       // Matching to PathData
       #parameterDefinition.directValues.cmdType := 3; // Circ Absolute
       #parameterDefinition.directValues.cmdParameters.circleParameters.circlePlane := 2; // XY
       #parameterDefinition.directValues.cmdParameters.circleParameters.pathChoice := 1; // neg rotation
       #parameterDefinition.directValues.cmdParameters.circleParameters.circMode := 3; // aux point is center relativ to start


     #G3:  // Circ CCW --> CircMode 1/2/3
       // Command name definition
       #parameterDefinition.parameterNameString := 'G';
       #parameterDefinition.parameterNameNumber := 3;

       // Properties
       #parameterDefinition.properties := "LKINLANG_MOTION_CMD" + "LKINLANG_CMD_MODAL";
       #parameterDefinition.validCountPerLine := 1;

       // Conditions
       #tempConditionCounter := 1;
       #parameterDefinition.conditions[#tempConditionCounter].ParameterNumber := #G17;
       #parameterDefinition.conditions[#tempConditionCounter].Group := 20;
       #parameterDefinition.conditions[#tempConditionCounter].Mode := "LKINLANG_CONDITION_IN_PROGRAM"; // In program
       #tempConditionCounter += 1;
       #parameterDefinition.conditions[#tempConditionCounter].ParameterNumber := #G18;
       #parameterDefinition.conditions[#tempConditionCounter].Group := 20;
       #parameterDefinition.conditions[#tempConditionCounter].Mode := "LKINLANG_CONDITION_IN_PROGRAM"; // In program
       #tempConditionCounter += 1;
       #parameterDefinition.conditions[#tempConditionCounter].ParameterNumber := #G19;
       #parameterDefinition.conditions[#tempConditionCounter].Group := 20;
       #parameterDefinition.conditions[#tempConditionCounter].Mode := "LKINLANG_CONDITION_IN_PROGRAM"; // In program
       #tempConditionCounter += 1;
       #parameterDefinition.conditions[#tempConditionCounter].ParameterNumber := #F;
       #parameterDefinition.conditions[#tempConditionCounter].Group := 10;
       #parameterDefinition.conditions[#tempConditionCounter].Mode := "LKINLANG_CONDITION_IN_PROGRAM"; // In program

       // Priorities
       // PathChoice and CmdType are defined
       #parameterDefinition.priorities.cmdType := "LKINLANG_PRIO_DEFINED";
       #parameterDefinition.priorities.cmdParameters.circleParameters.pathChoice := "LKINLANG_PRIO_DEFINED";

       // CircMode and circPlane can be changed (G17,G18,G19 / AR,CR,I,J,K)
       #parameterDefinition.priorities.cmdParameters.circleParameters.circlePlane := "LKINLANG_PRIO_DEFAULT";
       #parameterDefinition.priorities.cmdParameters.circleParameters.circMode := "LKINLANG_PRIO_DEFAULT";

       // Matching to PathData
       #parameterDefinition.directValues.cmdType := 3;
       #parameterDefinition.directValues.cmdParameters.circleParameters.circlePlane := 2; // XY
       #parameterDefinition.directValues.cmdParameters.circleParameters.pathChoice := 0; // pos rotation
       #parameterDefinition.directValues.cmdParameters.circleParameters.circMode := 3; // aux point is center relativ to start

     #G5:  // Circ 3D --> CircMode 0 
       // Command name definition
       #parameterDefinition.parameterNameString := 'G';
       #parameterDefinition.parameterNameNumber := 5;

       // Properties
       #parameterDefinition.properties := "LKINLANG_MOTION_CMD" + "LKINLANG_CMD_MODAL";
       #parameterDefinition.validCountPerLine := 1;

       // Conditions
       #tempConditionCounter := 1;
       #parameterDefinition.conditions[#tempConditionCounter].ParameterNumber := #F;
       #parameterDefinition.conditions[#tempConditionCounter].Group := 10;
       #parameterDefinition.conditions[#tempConditionCounter].Mode := "LKINLANG_CONDITION_IN_PROGRAM"; // In program

       // Priorities
       // CmdType and CircMode are defined 
       #parameterDefinition.priorities.cmdType := "LKINLANG_PRIO_DEFINED";
       #parameterDefinition.priorities.cmdParameters.circleParameters.circMode := "LKINLANG_PRIO_DEFINED";

       // Matching to PathData
       #parameterDefinition.directValues.cmdType := 3;
       #parameterDefinition.directValues.cmdParameters.circleParameters.circMode := 0; // aux point is on circ line


     #G4: // Wait time
       // Command name definition
       #parameterDefinition.parameterNameString := 'G';
       #parameterDefinition.parameterNameNumber := 4;

       // Properties
       #parameterDefinition.properties := 16#0;//"LKINLANG_MOTION_CMD";
       #parameterDefinition.validCountPerLine := 1;

       // Conditions
       #tempConditionCounter := 1;
       #parameterDefinition.conditions[#tempConditionCounter].ParameterNumber := #P;
       #parameterDefinition.conditions[#tempConditionCounter].Group := 30;
       #parameterDefinition.conditions[#tempConditionCounter].Mode := "LKINLANG_CONDITION_IN_LINE"; // In line

       #tempConditionCounter += 1;
       #parameterDefinition.conditions[#tempConditionCounter].ParameterNumber := #F;
       #parameterDefinition.conditions[#tempConditionCounter].Group := 30;
       #parameterDefinition.conditions[#tempConditionCounter].Mode := "LKINLANG_CONDITION_IN_LINE"; // In line

       // Properties
       #parameterDefinition.priorities.cmdType := "LKINLANG_PRIO_DEFINED";

       // Matching to PathData
       #parameterDefinition.directValues.cmdType := 100;

     #P: // WaitTime, same as F?
       // Command name definition
       #parameterDefinition.parameterNameString := 'P';
       #parameterDefinition.parameterNameNumber := -1;

       // Properties
       #parameterDefinition.properties := "LKINLANG_EQUATION";
       #parameterDefinition.validCountPerLine := 1;

       // Priorities
       #parameterDefinition.priorities.cmdParameters.pathDynamics.velocity := "LKINLANG_PRIO_DEFINED";

       // Matching to PathData
       #parameterDefinition.followingValues[1].cmdParameters.pathDynamics.velocity := TRUE;


     #G40: // Tool off
       // Command name definition
       #parameterDefinition.parameterNameString := 'G';
       #parameterDefinition.parameterNameNumber := 40;

       // Properties
       #parameterDefinition.properties := 16#0;//"LKINLANG_MOTION_CMD";

       // Priorities
       #parameterDefinition.priorities.cmdType := "LKINLANG_PRIO_DEFINED";

       // Matching to PathData
       #parameterDefinition.directValues.cmdType := 40;

     #G41: // Tool left
       // Command name definition
       #parameterDefinition.parameterNameString := 'G';
       #parameterDefinition.parameterNameNumber := 41;

       // Properties
       #parameterDefinition.properties := 16#0;//"LKINLANG_MOTION_CMD";

       // Priorities
       #parameterDefinition.priorities.cmdType := "LKINLANG_PRIO_DEFINED";

       // Matching to PathData
       #parameterDefinition.directValues.cmdType := 41;

       // Conditions
       #tempConditionCounter := 1;
       #parameterDefinition.conditions[#tempConditionCounter].ParameterNumber := #T;
       #parameterDefinition.conditions[#tempConditionCounter].Group := 40;
       #parameterDefinition.conditions[#tempConditionCounter].Mode := "LKINLANG_CONDITION_IN_PROGRAM";
       #tempConditionCounter += 1;
       #parameterDefinition.conditions[#tempConditionCounter].ParameterNumber := #G17;
       #parameterDefinition.conditions[#tempConditionCounter].Group := 20;
       #parameterDefinition.conditions[#tempConditionCounter].Mode := "LKINLANG_CONDITION_IN_PROGRAM"; // In program
       #tempConditionCounter += 1;
       #parameterDefinition.conditions[#tempConditionCounter].ParameterNumber := #G18;
       #parameterDefinition.conditions[#tempConditionCounter].Group := 20;
       #parameterDefinition.conditions[#tempConditionCounter].Mode := "LKINLANG_CONDITION_IN_PROGRAM"; // In program
       #tempConditionCounter += 1;
       #parameterDefinition.conditions[#tempConditionCounter].ParameterNumber := #G19;
       #parameterDefinition.conditions[#tempConditionCounter].Group := 20;
       #parameterDefinition.conditions[#tempConditionCounter].Mode := "LKINLANG_CONDITION_IN_PROGRAM"; // In program

     #G42: // Tool right
       // Command name definition
       #parameterDefinition.parameterNameString := 'G';
       #parameterDefinition.parameterNameNumber := 42;

       // Properties
       #parameterDefinition.properties := 16#0; //"LKINLANG_MOTION_CMD";

       // Priorities
       #parameterDefinition.priorities.cmdType := "LKINLANG_PRIO_DEFINED";

       // Matching to PathData
       #parameterDefinition.directValues.cmdType := 42;

       // Conditions
       #tempConditionCounter := 1;
       #parameterDefinition.conditions[#tempConditionCounter].ParameterNumber := #T;
       #parameterDefinition.conditions[#tempConditionCounter].Group := 40;
       #parameterDefinition.conditions[#tempConditionCounter].Mode := "LKINLANG_CONDITION_IN_PROGRAM";
       #tempConditionCounter += 1;
       #parameterDefinition.conditions[#tempConditionCounter].ParameterNumber := #G17;
       #parameterDefinition.conditions[#tempConditionCounter].Group := 20;
       #parameterDefinition.conditions[#tempConditionCounter].Mode := "LKINLANG_CONDITION_IN_PROGRAM"; // In program
       #tempConditionCounter += 1;
       #parameterDefinition.conditions[#tempConditionCounter].ParameterNumber := #G18;
       #parameterDefinition.conditions[#tempConditionCounter].Group := 20;
       #parameterDefinition.conditions[#tempConditionCounter].Mode := "LKINLANG_CONDITION_IN_PROGRAM"; // In program
       #tempConditionCounter += 1;
       #parameterDefinition.conditions[#tempConditionCounter].ParameterNumber := #G19;
       #parameterDefinition.conditions[#tempConditionCounter].Group := 20;
       #parameterDefinition.conditions[#tempConditionCounter].Mode := "LKINLANG_CONDITION_IN_PROGRAM"; // In program

     #T: // Tool selection
       // Command name definition
       #parameterDefinition.parameterNameString := 'T';
       #parameterDefinition.parameterNameNumber := -1;

       #parameterDefinition.validCountPerLine := 1;

       // Properties
       #parameterDefinition.properties := "LKINLANG_PRG_MODAL";

       // Matching to PathData
       #parameterDefinition.priorities.cmdParameters.offsetParameters.offsetParaNo := "LKINLANG_PRIO_DEFINED";
       #parameterDefinition.followingValues[1].cmdParameters.offsetParameters.offsetParaNo := TRUE;


     #G17: // XY PathPlane
       // Command name definition
       #parameterDefinition.parameterNameString := 'G';
       #parameterDefinition.parameterNameNumber := 17;

       // Properties
       #parameterDefinition.properties := "LKINLANG_PRG_MODAL";

       // Matching to PathData
       #parameterDefinition.priorities.cmdParameters.circleParameters.circlePlane := "LKINLANG_PRIO_DEFINED";
       #parameterDefinition.directValues.cmdParameters.circleParameters.circlePlane := 2; // XY

       // Also set main path plane
       #parameterDefinition.priorities.cmdParameters.offsetParameters.mainPathPlane := "LKINLANG_PRIO_DEFINED";
       #parameterDefinition.directValues.cmdParameters.offsetParameters.mainPathPlane := 2; // XY

     #G18: // XZ PathPlane
       // Command name definition
       #parameterDefinition.parameterNameString := 'G';
       #parameterDefinition.parameterNameNumber := 18;

       // Properties
       #parameterDefinition.properties := "LKINLANG_PRG_MODAL";

       // Matching to PathData
       #parameterDefinition.priorities.cmdParameters.circleParameters.circlePlane := "LKINLANG_PRIO_DEFINED";
       #parameterDefinition.directValues.cmdParameters.circleParameters.circlePlane := 0; // XZ

       // Also set main path plane
       #parameterDefinition.priorities.cmdParameters.offsetParameters.mainPathPlane := "LKINLANG_PRIO_DEFINED";
       #parameterDefinition.directValues.cmdParameters.offsetParameters.mainPathPlane := 0; // XZ

     #G19: //YZ PathPlane
       // Command name definition
       #parameterDefinition.parameterNameString := 'G';
       #parameterDefinition.parameterNameNumber := 19;

       // Properties
       #parameterDefinition.properties := "LKINLANG_PRG_MODAL";

       // Matching to PathData
       #parameterDefinition.priorities.cmdParameters.circleParameters.circlePlane := "LKINLANG_PRIO_DEFINED";
       #parameterDefinition.directValues.cmdParameters.circleParameters.circlePlane := 1; // YZ

       // Also set main path plane
       #parameterDefinition.priorities.cmdParameters.offsetParameters.mainPathPlane := "LKINLANG_PRIO_DEFINED";
       #parameterDefinition.directValues.cmdParameters.offsetParameters.mainPathPlane := 1; // YZ

     #G640:
       // Command name definition
       #parameterDefinition.parameterNameString := 'G';
       #parameterDefinition.parameterNameNumber := 640;

       // Properties
       #parameterDefinition.properties := "LKINLANG_PRG_MODAL";

       // Matching to PathData
       #parameterDefinition.priorities.cmdParameters.bufferMode := "LKINLANG_PRIO_DEFINED";
       #parameterDefinition.directValues.cmdParameters.bufferMode := 1; // Standstill

       #parameterDefinition.priorities.cmdParameters.transitionParameters[1] := "LKINLANG_PRIO_DEFINED";
       #parameterDefinition.directValues.cmdParameters.transitionParameters[1] := 0.0; // Standstill

     #G641:
       // Command name definition
       #parameterDefinition.parameterNameString := 'G';
       #parameterDefinition.parameterNameNumber := 641;

       // Properties
       #parameterDefinition.properties := "LKINLANG_PRG_MODAL";

       // Conditions
       #tempConditionCounter := 1;
       #parameterDefinition.conditions[#tempConditionCounter].ParameterNumber := #BR;
       #parameterDefinition.conditions[#tempConditionCounter].Group := 50;
       #parameterDefinition.conditions[#tempConditionCounter].Mode := "LKINLANG_CONDITION_IN_LINE"; // In line

       // Matching to PathData
       #parameterDefinition.priorities.cmdParameters.bufferMode := "LKINLANG_PRIO_DEFINED";
       #parameterDefinition.directValues.cmdParameters.bufferMode := #parameterDefaults.transitionVelocityMode;

     #G90:
       // Command name definition
       #parameterDefinition.parameterNameString := 'G';
       #parameterDefinition.parameterNameNumber := 90;

       // Properties
       #parameterDefinition.properties := "LKINLANG_PRG_MODAL" + "LKINLANG_ABSOLUTE_POSITION";


     #G91:
       // Command name definition
       #parameterDefinition.parameterNameString := 'G';
       #parameterDefinition.parameterNameNumber := 91;

       // Properties
       #parameterDefinition.properties := "LKINLANG_PRG_MODAL" + "LKINLANG_RELATIVE_POSITION";

     #G54: // Select OCS 1
       // Command name definition
       #parameterDefinition.parameterNameString := 'G';
       #parameterDefinition.parameterNameNumber := 54;

       // Properties
       #parameterDefinition.properties := "LKINLANG_PRG_MODAL" + "LKINLANG_CHECK_LIMITS";

       // Matching to PathData
       #parameterDefinition.priorities.cmdCoordinates.coordSystem := "LKINLANG_PRIO_DEFINED";
       #parameterDefinition.directValues.cmdCoordinates.coordSystem := 1; // OCS1


     #G55: // Select OCS 2
       // Command name definition
       #parameterDefinition.parameterNameString := 'G';
       #parameterDefinition.parameterNameNumber := 55;

       // Properties
       #parameterDefinition.properties := "LKINLANG_PRG_MODAL" + "LKINLANG_CHECK_LIMITS";

       // Matching to PathData
       #parameterDefinition.priorities.cmdCoordinates.coordSystem := "LKINLANG_PRIO_DEFINED";
       #parameterDefinition.directValues.cmdCoordinates.coordSystem := 2; // OCS2


     #G56: // Select OCS 3
       // Command name definition
       #parameterDefinition.parameterNameString := 'G';
       #parameterDefinition.parameterNameNumber := 56;

       // Properties
       #parameterDefinition.properties := "LKINLANG_PRG_MODAL" + "LKINLANG_CHECK_LIMITS";

       // Matching to PathData
       #parameterDefinition.priorities.cmdCoordinates.coordSystem := "LKINLANG_PRIO_DEFINED";
       #parameterDefinition.directValues.cmdCoordinates.coordSystem := 3; // OCS3


     #G500: // Select WCS
       // Command name definition
       #parameterDefinition.parameterNameString := 'G';
       #parameterDefinition.parameterNameNumber := 500;

       // Properties
       #parameterDefinition.properties := "LKINLANG_PRG_MODAL" + "LKINLANG_CHECK_LIMITS";

       // Matching to PathData
       #parameterDefinition.priorities.cmdCoordinates.coordSystem := "LKINLANG_PRIO_DEFINED";
       #parameterDefinition.directValues.cmdCoordinates.coordSystem := 0; // WCS


       // Gerneral Parameters (170 - 199)
       // ===========================================================
     #X:
       #parameterDefinition.parameterNameString := 'X';
       #parameterDefinition.parameterNameNumber := -1;
       #parameterDefinition.properties := "LKINLANG_CHECK_LIMITS" + "LKINLANG_EQUATION";
       #parameterDefinition.priorities.cmdCoordinates.cartesianPosition.x := "LKINLANG_PRIO_DEFINED";
       #parameterDefinition.followingValues[1].cmdCoordinates.cartesianPosition.x := true;

     #Y:
       #parameterDefinition.parameterNameString := 'Y';
       #parameterDefinition.parameterNameNumber := -1;
       #parameterDefinition.properties := "LKINLANG_CHECK_LIMITS" + "LKINLANG_EQUATION";
       #parameterDefinition.priorities.cmdCoordinates.cartesianPosition.y := "LKINLANG_PRIO_DEFINED";
       #parameterDefinition.followingValues[1].cmdCoordinates.cartesianPosition.y := true;

     #Z:
       #parameterDefinition.parameterNameString := 'Z';
       #parameterDefinition.parameterNameNumber := -1;
       #parameterDefinition.properties := "LKINLANG_CHECK_LIMITS" + "LKINLANG_EQUATION";
       #parameterDefinition.priorities.cmdCoordinates.cartesianPosition.z := "LKINLANG_PRIO_DEFINED";
       #parameterDefinition.followingValues[1].cmdCoordinates.cartesianPosition.z := true;

     #A:
       #parameterDefinition.parameterNameString := 'A';
       #parameterDefinition.parameterNameNumber := -1;
       #parameterDefinition.properties := "LKINLANG_CHECK_LIMITS" + "LKINLANG_EQUATION";
       #parameterDefinition.priorities.cmdCoordinates.cartesianPosition.a := "LKINLANG_PRIO_DEFINED";
       #parameterDefinition.followingValues[1].cmdCoordinates.cartesianPosition.a := true;

       // Orientation direction
       #parameterDefinition.directValues.cmdParameters.orientationDirection := #parameterDefaults.orientationDirection;
       #parameterDefinition.directValues.cmdParameters.orientationDirection := "LKINLANG_PRIO_DEFAULT";

     #F:
       #parameterDefinition.parameterNameString := 'F';
       #parameterDefinition.parameterNameNumber := -1;
       #parameterDefinition.properties := "LKINLANG_PRG_MODAL" + "LKINLANG_CHECK_LIMITS" + "LKINLANG_EQUATION";
       #parameterDefinition.priorities.cmdParameters.pathDynamics.velocity := "LKINLANG_PRIO_DEFINED";
       #parameterDefinition.followingValues[1].cmdParameters.pathDynamics.velocity := TRUE;

     #ACC:
       #parameterDefinition.parameterNameString := 'ACC';
       #parameterDefinition.parameterNameNumber := -1;
       #parameterDefinition.properties := "LKINLANG_PRG_MODAL" + "LKINLANG_CHECK_LIMITS" + "LKINLANG_EQUATION";
       #parameterDefinition.priorities.cmdParameters.pathDynamics.acceleration := "LKINLANG_PRIO_DEFINED";
       #parameterDefinition.followingValues[1].cmdParameters.pathDynamics.acceleration := TRUE;

     #DEC:
       #parameterDefinition.parameterNameString := 'DEC';
       #parameterDefinition.parameterNameNumber := -1;
       #parameterDefinition.properties := "LKINLANG_PRG_MODAL" + "LKINLANG_CHECK_LIMITS" + "LKINLANG_EQUATION";
       #parameterDefinition.priorities.cmdParameters.pathDynamics.deceleration := "LKINLANG_PRIO_DEFINED";
       #parameterDefinition.followingValues[1].cmdParameters.pathDynamics.deceleration := TRUE;

     #JERK:
       #parameterDefinition.parameterNameString := 'JERK';
       #parameterDefinition.parameterNameNumber := -1;
       #parameterDefinition.properties := "LKINLANG_PRG_MODAL" + "LKINLANG_CHECK_LIMITS" + "LKINLANG_EQUATION";
       #parameterDefinition.priorities.cmdParameters.pathDynamics.jerk := "LKINLANG_PRIO_DEFINED";
       #parameterDefinition.followingValues[1].cmdParameters.pathDynamics.jerk := TRUE;


     #I:
       // Command name definition
       #parameterDefinition.parameterNameString := 'I';
       #parameterDefinition.parameterNameNumber := -1;

       // Properties
       #parameterDefinition.properties := "LKINLANG_EQUATION";

       // Matching to PathData
       #parameterDefinition.priorities.cmdParameters.circleParameters.auxPoint[1] := "LKINLANG_PRIO_DEFINED";
       #parameterDefinition.followingValues[1].cmdParameters.circleParameters.auxPoint[1] := TRUE;

     #J:
       // Command name definition
       #parameterDefinition.parameterNameString := 'J';
       #parameterDefinition.parameterNameNumber := -1;

       // Properties
       #parameterDefinition.properties := "LKINLANG_EQUATION";

       // Matching to PathData
       #parameterDefinition.priorities.cmdParameters.circleParameters.auxPoint[2] := "LKINLANG_PRIO_DEFINED";
       #parameterDefinition.followingValues[1].cmdParameters.circleParameters.auxPoint[2] := TRUE;

     #K:
       // Command name definition
       #parameterDefinition.parameterNameString := 'K';
       #parameterDefinition.parameterNameNumber := -1;

       // Properties
       #parameterDefinition.properties := "LKINLANG_EQUATION";

       // Matching to PathData
       #parameterDefinition.priorities.cmdParameters.circleParameters.auxPoint[3] := "LKINLANG_PRIO_DEFINED";
       #parameterDefinition.followingValues[1].cmdParameters.circleParameters.auxPoint[3] := TRUE;

     #AR:
       // Command name definition
       #parameterDefinition.parameterNameString := 'AR';
       #parameterDefinition.parameterNameNumber := -1;

       // Properties
       #parameterDefinition.properties := "LKINLANG_EQUATION";

       // Conditions
       #tempConditionCounter := 1;
       #parameterDefinition.conditions[#tempConditionCounter].ParameterNumber := #I;
       #parameterDefinition.conditions[#tempConditionCounter].Group := 60;
       #parameterDefinition.conditions[#tempConditionCounter].Mode := "LKINLANG_CONDITION_IN_LINE"; // In Line
       #tempConditionCounter += 1; 
       #parameterDefinition.conditions[#tempConditionCounter].ParameterNumber := #J;
       #parameterDefinition.conditions[#tempConditionCounter].Group := 60;
       #parameterDefinition.conditions[#tempConditionCounter].Mode := "LKINLANG_CONDITION_IN_LINE"; // In Line
       #tempConditionCounter += 1;
       #parameterDefinition.conditions[#tempConditionCounter].ParameterNumber := #K;
       #parameterDefinition.conditions[#tempConditionCounter].Group := 60;
       #parameterDefinition.conditions[#tempConditionCounter].Mode := "LKINLANG_CONDITION_IN_LINE"; // In Line

       // Matching to PathData
       #parameterDefinition.priorities.cmdParameters.circleParameters.arc := "LKINLANG_PRIO_DEFINED";
       #parameterDefinition.followingValues[1].cmdParameters.circleParameters.arc := TRUE;
       #parameterDefinition.priorities.cmdParameters.circleParameters.circMode := "LKINLANG_PRIO_DEFINED";
       #parameterDefinition.directValues.cmdParameters.circleParameters.circMode := 1;

     #CR:
       // Command name definition
       #parameterDefinition.parameterNameString := 'CR';
       #parameterDefinition.parameterNameNumber := -1;

       // Properties
       #parameterDefinition.properties := "LKINLANG_EQUATION";

       // Conditions
       #tempConditionCounter := 1;
       #parameterDefinition.conditions[#tempConditionCounter].ParameterNumber := #X;
       #parameterDefinition.conditions[#tempConditionCounter].Group := 70;
       #parameterDefinition.conditions[#tempConditionCounter].Mode := "LKINLANG_CONDITION_IN_LINE"; // In Line
       #tempConditionCounter += 1;
       #parameterDefinition.conditions[#tempConditionCounter].ParameterNumber := #Y;
       #parameterDefinition.conditions[#tempConditionCounter].Group := 70;
       #parameterDefinition.conditions[#tempConditionCounter].Mode := "LKINLANG_CONDITION_IN_LINE"; // In Line
       #tempConditionCounter += 1;
       #parameterDefinition.conditions[#tempConditionCounter].ParameterNumber := #Z;
       #parameterDefinition.conditions[#tempConditionCounter].Group := 70;
       #parameterDefinition.conditions[#tempConditionCounter].Mode := "LKINLANG_CONDITION_IN_LINE"; // In Line

       // Matching to PathData
       #parameterDefinition.priorities.cmdParameters.circleParameters.radius := "LKINLANG_PRIO_DEFINED";
       #parameterDefinition.followingValues[1].cmdParameters.circleParameters.radius := TRUE;
       #parameterDefinition.priorities.cmdParameters.circleParameters.circMode := "LKINLANG_PRIO_DEFINED";
       #parameterDefinition.directValues.cmdParameters.circleParameters.circMode := 2;

     #M:
       // Command name definition
       #parameterDefinition.parameterNameString := 'M';
       #parameterDefinition.parameterNameNumber := -1;

       #parameterDefinition.validCountPerLine := "LKINCTRL_NO_OF_CMD_SETFLAGS";

       // Properties
       #parameterDefinition.properties := "LKINLANG_CHECK_LIMITS";

       // Matching to PathData
       #parameterDefinition.priorities.setFlags.flag := "LKINLANG_PRIO_DEFINED";
       #parameterDefinition.priorities.setFlags.flagMode := "LKINLANG_PRIO_DEFINED";
       #parameterDefinition.priorities.setFlags.remainingDistance := "LKINLANG_PRIO_DEFINED";
       #parameterDefinition.followingValues[1].setFlags.flag := TRUE;
       #parameterDefinition.followingValues[2].setFlags.flagMode := TRUE;
       #parameterDefinition.followingValues[3].setFlags.remainingDistance := TRUE;

     #H:
       // Command name definition
       #parameterDefinition.parameterNameString := 'H';
       #parameterDefinition.parameterNameNumber := -1;

       #parameterDefinition.validCountPerLine := "LKINCTRL_NO_OF_CMD_SETFLAGS";

       // Properties
       #parameterDefinition.properties := "LKINLANG_CHECK_LIMITS" + "LKINLANG_EQUATION";

       // Matching to PathData
       #parameterDefinition.priorities.valueFlags.flag := "LKINLANG_PRIO_DEFINED";
       #parameterDefinition.priorities.valueFlags.value := "LKINLANG_PRIO_DEFINED";
       #parameterDefinition.priorities.valueFlags.flagMode := "LKINLANG_PRIO_DEFINED";
       #parameterDefinition.priorities.valueFlags.remainingDistance := "LKINLANG_PRIO_DEFINED";
       #parameterDefinition.followingValues[1].valueFlags.flag := TRUE;
       #parameterDefinition.followingValues[2].valueFlags.value := TRUE;
       #parameterDefinition.followingValues[3].valueFlags.flagMode := TRUE;
       #parameterDefinition.followingValues[4].valueFlags.remainingDistance := TRUE;

     #BR:
       // Command name definition
       #parameterDefinition.parameterNameString := 'BR';
       #parameterDefinition.parameterNameNumber := -1;

       // Properties
       #parameterDefinition.properties := "LKINLANG_PRG_MODAL" + "LKINLANG_EQUATION";

       // Matching to PathData
       #parameterDefinition.priorities.cmdParameters.transitionParameters[1] := "LKINLANG_PRIO_DEFINED";
       #parameterDefinition.followingValues[1].cmdParameters.transitionParameters[1] := TRUE;

     #M30:
       // Command name definition
       #parameterDefinition.parameterNameString := 'M';
       #parameterDefinition.parameterNameNumber := 30;

       #parameterDefinition.validCountPerLine := 1;

       // Properties
       #parameterDefinition.properties := "LKINLANG_MOTION_CMD";
       #parameterDefinition.priorities.cmdType := "LKINLANG_PRIO_DEFINED";

       // Matching to PathData
       #parameterDefinition.directValues.cmdType := -1;
     ELSE
       // invalid case number
       #parameterNo := -2;

   END_CASE;
END_FUNCTION

FUNCTION "LKinLang_UserDefinedGCode" : Void   // FC35453, SCL
TITLE = LKinLang_LangPackageGCode
{ S7_Optimized_Access := 'TRUE' }
AUTHOR : tech.team.motioncontrol@siemens.com
FAMILY : LKinLang
VERSION : 1.1
// Language definition package for user defined GCode
   VAR_IN_OUT
      parameterNo : Int;   // Parameter number
      parameterDefinition : "LKinLang_typeParameterDefinition";   // Found parameter definition
      parameterDefaults : "LKinLang_typeGCodeDefaults";   // Parameter defaults
   END_VAR
   VAR_TEMP
      tempConditionCounter : Int;
   END_VAR
   VAR CONSTANT
      G0 : DInt := 100;   // Fast Lin
      G1 : DInt := 101;   // Lin
      G2 : DInt := 102;   // Circ CW
      G3 : DInt := 103;   // Circ CCW
      G5 : DInt := 105;   // Circ 3D
      G4 : DInt := 104;   // WaitTime
      P : DInt := 110;   // Period for WaitTime
      G17 : DInt := 120;   // XY Plane
      G18 : DInt := 121;   // ZX Plane
      G19 : DInt := 122;   // YZ Plane
      G640 : DInt := 130;   // Geometry blending off
      G641 : DInt := 131;   // Geometry blending with high velocity
      G642 : DInt := 132;   // Geometry blending with low velocity
      G90 : DInt := 150;   // Absolute Position
      G91 : DInt := 151;   // Relativ Position
      G54 : DInt := 152;   // Select OCS1
      G55 : DInt := 153;   // Select OCS2
      G56 : DInt := 154;   // Select OCS3
      G500 : DInt := 155;   // Select WCS
      T : DInt := 160;   // Tool selection
      G40 : DInt := 161;   // Tool off
      G41 : DInt := 162;   // Tool left
      G42 : DInt := 163;   // Tool right
      X : DInt := 170;   // X pos
      Y : DInt := 171;   // Y pos
      Z : DInt := 172;   // Z pos
      "A" : DInt := 173;   // Orientation
      F : DInt := 174;   // Velocity
      ACC : DInt := 175;   // Acceleration
      DEC : DInt := 176;   // Deceleration
      JERK : DInt := 177;   // Jerk
      CR : DInt := 178;   // Circle Radius
      I : DInt := 179;   // Circ Point
      J : DInt := 180;   // Circ Point
      K : DInt := 181;   // Circ Point
      AR : DInt := 182;   // Arc
      BR : DInt := 183;   // Transition Parameter
      "M" : DInt := 190;   // Flag
      M30 : DInt := 199;   // End of PRG
   END_VAR
BEGIN
   //==========================================================================================
   // SIEMENS AG
   // (c)Copyright 2019 All Rights Reserved
   //------------------------------------------------------------------------------------------
   // Library: LKinLang
   // Tested with: S7-1517T-3 PN/DP
   // Engineering: TIA Portal V15
   // Restrictions: ---
   // Requirements: S7-1500T FW 2.5
   // Functionality: LKinLang_UserDefinedGCode
   // Language definition package for user defined GCode
   // 
   // Support: tech.team.motioncontrol@siemens.com
   // Note: Parameter comments are only available in language 'English (United States)'
   //------------------------------------------------------------------------------------------
   // Change log table:
   // Version    Date          Expert in charge    Changes applied
   // 01.00.00   28.05.2019    FR                  First created version
   //===========================================================================================
   //
   //  Group Parameter 
   //  10:   F
   //        
   //  20:   G17
   //        G18
   //        G19
   //        
   //  30:   F
   //        P
   //        
   //  40:   T
   //
   //  50:   BR
   //  
   //  60:   I
   //        J
   //        K
   //
   //  70:   X
   //        Y
   //        Z


   CASE #parameterNo OF
       // User defined commands for GCode.
       // Here you can define up to 100 commands.
       // It is possible to overload predefined GCode commands.
       // Or define own commands.
       // Some example are already programmed.
       // ------------------------------
     1:
       // ========================================================================================================
       // End of program
       // ========================================================================================================
       // Instead of M30, END is also possible
       // ========================================================================================================
       // Parameter name definition
       #parameterDefinition.parameterNameString := 'END';
       #parameterDefinition.parameterNameNumber := -1;

       // Matching to PathData
       #parameterDefinition.directValues.cmdType := -1;

       // Priorities
       #parameterDefinition.priorities.cmdType := "LKINLANG_PRIO_DEFINED";

       // Properties
       #parameterDefinition.properties := "LKINLANG_MOTION_CMD";

       // Valid counts per line
       #parameterDefinition.validCountPerLine := 1;
       // ========================================================================================================

     2:
       // ========================================================================================================
       // Gripper control ON
       // ========================================================================================================
       // This is an example for an defined "Gripper" parameter
       // 'GRIPPER_ON' sets Flag 1 with Flagmode 11
       // ========================================================================================================
       // Parameter name definition
       #parameterDefinition.parameterNameString := 'GRIPPER_ON';
       #parameterDefinition.parameterNameNumber := -1;

       // Matching to PathData
       #parameterDefinition.directValues.setFlags[1].flag := 1;
       #parameterDefinition.directValues.setFlags[1].flagMode := 11;

       // Priorities
       #parameterDefinition.priorities.setFlags.flag := "LKINLANG_PRIO_DEFINED";
       #parameterDefinition.priorities.setFlags.flagMode := "LKINLANG_PRIO_DEFINED";

       // Properties
       #parameterDefinition.properties := 16#0;

       // Valid counts per line
       #parameterDefinition.validCountPerLine := 1;
       // ========================================================================================================

     3:
       // ========================================================================================================
       // Gripper control OFF
       // ========================================================================================================
       // This is an example for an defined "Gripper" parameter
       // 'GRIPPER_OFF' resets Flag 1 with Flagmode 13
       // ========================================================================================================
       // Parameter name definition
       #parameterDefinition.parameterNameString := 'GRIPPER_OFF';
       #parameterDefinition.parameterNameNumber := -1;

       // Matching to PathData
       #parameterDefinition.directValues.setFlags[1].flag := 1;
       #parameterDefinition.directValues.setFlags[1].flagMode := 13;

       // Priorities
       #parameterDefinition.priorities.setFlags.flag := "LKINLANG_PRIO_DEFINED";
       #parameterDefinition.priorities.setFlags.flagMode := "LKINLANG_PRIO_DEFINED";

       // Properties
       #parameterDefinition.properties := 16#0;

       // Valid counts per line
       #parameterDefinition.validCountPerLine := 1;
       // ========================================================================================================

     4: 
       // ========================================================================================================
       // Point name
       // ========================================================================================================
       // Use 'Nxx' as point name in the PathData
       // --> Only numbers possible
       // ========================================================================================================
       // Parameter name definition
       #parameterDefinition.parameterNameString := 'N';
       #parameterDefinition.parameterNameNumber := -1;

       // Matching to PathData
       #parameterDefinition.followingValues[1].cmdName := TRUE;

       // Priorities
       #parameterDefinition.priorities.cmdName := "LKINLANG_PRIO_DEFINED";

       // Properties
       #parameterDefinition.properties := 16#0;

       // Valid counts per line
       #parameterDefinition.validCountPerLine := 1;
       // ========================================================================================================

     5:
       // ========================================================================================================
       // Blending with low velocity
       // ========================================================================================================
       // Parameter name definition
       #parameterDefinition.parameterNameString := 'G';
       #parameterDefinition.parameterNameNumber := 642;

       // Matching to PathData
       #parameterDefinition.directValues.cmdParameters.bufferMode := 2; // Blending with low velocity

       // Priorites
       #parameterDefinition.priorities.cmdParameters.bufferMode := "LKINLANG_PRIO_DEFINED";

       // Properties
       #parameterDefinition.properties := "LKINLANG_PRG_MODAL";

       // Conditions
       #tempConditionCounter := 1;
       #parameterDefinition.conditions[#tempConditionCounter].ParameterNumber := #BR;
       #parameterDefinition.conditions[#tempConditionCounter].Group := 50;
       #parameterDefinition.conditions[#tempConditionCounter].Mode := "LKINLANG_CONDITION_IN_LINE"; // "BR" must be written in the same line

       // Valid counts per line
       #parameterDefinition.validCountPerLine := 1;
       // ========================================================================================================

     ELSE
       // invalid case number
       #parameterNo := -2;
   END_CASE;
END_FUNCTION

// folder: LKinLang_Blocks/LKinLang_LanguageDefinition/LKinLang_LangPackUser

FUNCTION "LKinLang_LangPackageUser" : Void   // FC35487, SCL
TITLE = LKinLang_LangPackageUser
{ S7_Optimized_Access := 'TRUE' }
AUTHOR : tech.team.motioncontrol@siemens.com
FAMILY : LKinLang
VERSION : 1.1
// Language definition package for a user defined language
   VAR_IN_OUT
      parameterNo : Int;   // Parameter number
      parameterDefinition : "LKinLang_typeParameterDefinition";   // Found parameter definition / Found command definition
      parameterDefaults : "LKinLang_typeUserDefinedDefaults";   // Parameter defaults
   END_VAR
   VAR_TEMP
      tempConditionCounter : Int;   // Temporary counter
   END_VAR
   VAR CONSTANT
      LIN : DInt := 1;   // Fast Lin
      VEL : DInt := 2;   // Velocity / Circ CW
      BLEND : DInt := 3;   // Blending
      RADIUS : DInt := 4;   // Blending radius
      X : DInt := 5;   // X pos
      Y : DInt := 6;   // Y pos
      Z : DInt := 7;   // Z pos
      END : DInt := 8;   // End of PRG
   END_VAR
BEGIN
   //==========================================================================================
   // SIEMENS AG
   // (c)Copyright 2019 All Rights Reserved
   //------------------------------------------------------------------------------------------
   // Library: LKinLang
   // Tested with: S7-1517T-3 PN/DP
   // Engineering: TIA Portal V15
   // Restrictions: ---
   // Requirements: S7-1500T FW 2.5
   // Functionality: LKinLang_LangPackageUser
   // Language definition package for completly user defined language
   // 
   // Support: tech.team.motioncontrol@siemens.com
   // Note: Parameter comments are only available in language 'English (United States)'
   //------------------------------------------------------------------------------------------
   // Change log table:
   // Version    Date          Expert in charge    Changes applied
   // 01.00.00   28.05.2019    FR                  First created version
   //===========================================================================================
   //
   //  Group Parameter 
   //  10:   R
   //        

   CASE #parameterNo OF
       // ========================================================================================================
       // Motion Parameters
       // ========================================================================================================
     #LIN:
       // ========================================================================================================
       // Linear movement
       // ========================================================================================================
       // Definition of linear movement (PathData: cmdType = 1) with default velocity
       // Parameter name is defined by parameterNameString and parameterNameNumber
       // ParameterNameString = LIN
       // ParameterNameNumber = -1 --> irrelevant
       // ==> Program line is searched for "LIN"

       // If "LIN" was found, set the defined values in the connected PathData.
       // The values are defined as "DirectValues" because the value to set is directly written here in this FC
       // Command type (cmdType)
       // #parameterDefinition.directValues.cmdType := 1;
       // --> Set the cmdType to 1
       // 
       // Velocity
       // #parameterDefinition.directValues.cmdParameters.pathDynamics.velocity := #parameterDefaults.velocityLin;
       // --> Set the path velocity to the value set in the variable #parameterDefaults.velocityLin
       // 
       // Parameter Priorities:
       // ----------
       // The priorities define if a value can be overwritten by another parameter.
       // e.g. The velocity is set with prio "LKINLANG_PRIO_DEFAULT", this means the velocity can be overwritten by every other parameter
       // which has a velocity prio higher than "LKINLANG_PRIO_DEFAULT".
       // 
       // The priorities are as followed:
       // Lowest:  "LKINLANG_PRIO_UNRELEVANT"
       //          "LKINLANG_PRIO_DEFAULT" 
       //          "LKINLANG_PRIO_DEFINED"
       // Highest: "LKINLANG_PRIO_CONSTANT"
       // 
       //
       // Parameter properties:
       // ----------
       // Properties can be used to define parameters as motion command or as modal.
       // To do so, add all properties you want to have.
       // e.g. LIN is a motion command therfore the property "LKINLANG_MOTION_CMD" is set.
       // Also it shall be modal until the motion command changes, so the property "LKINLANG_CMD_MODAL" is set.
       // 
       //
       // The properties are as followed:
       // ----------
       // "LKINLANG_MOTION_CMD" --> Is motion command
       // "LKINLANG_ABSOLUTE_POSITION" --> Switch to absolute positioning 
       // "LKINLANG_RELATIVE_POSITION" --> Switch to relative positioning
       // "LKINLANG_CMD_MODAL" --> Modal until change of motion cmd
       // "LKINLANG_PRG_MODAL" --> Modal in program until overwritten
       // "LKINLANG_CHECK_LIMITS" --> Check the limits for written elements (e.g. cmdType > -1 and < 101)
       // "LKINLANG_EQUATION" --> Mathematical expression allowed after parameter
       //
       // 
       // ValidCountPerLine:
       // ----------
       // This value defines how often the same parameter can occur in the same line.
       // The default setting is 1
       // 
       // Parameter name definition
       #parameterDefinition.parameterNameString := 'LIN';
       #parameterDefinition.parameterNameNumber := -1;

       // Matching to PathData
       #parameterDefinition.directValues.cmdType := 1;
       #parameterDefinition.directValues.cmdParameters.pathDynamics.velocity := #parameterDefaults.velocityLin;

       // Priorities
       #parameterDefinition.priorities.cmdType := "LKINLANG_PRIO_DEFINED";
       #parameterDefinition.priorities.cmdParameters.pathDynamics.velocity := "LKINLANG_PRIO_DEFAULT";

       // Properties
       #parameterDefinition.properties := "LKINLANG_MOTION_CMD" + "LKINLANG_CMD_MODAL";

       // Valid counts per line
       #parameterDefinition.validCountPerLine := 1;
       // ========================================================================================================


     #VEL:
       // ========================================================================================================
       // Path Velocity
       // ========================================================================================================
       // Definition of path velocity (PathData: cmdParameters.pathDynamics.velocity)
       // The parameter name is defined as "VEL"
       // 
       // If "VEL" was found, set the defined values in the connected PathData
       // The value is defined as "FollowingValue" because the value is not written here, but in the program line after this parameter
       // e.g. VEL=200 <-- 200 is taken as path velocity
       // To do this, set #parameterDefinition.followingValues[1].cmdParameters.pathDynamics.velocity := TRUE;
       // 
       // Also set the priority #parameterDefinition.priorities.cmdParameters.pathDynamics.velocity := "LKINLANG_PRIO_DEFINED";
       // 
       // Properties:
       // ----------
       // "LKINLANG_PRG_MODAL": Modal in program to save velocity value once set
       // "LKINLANG_EQUATION": Allow mathematical expressions (e.g. VEL=200+10)
       //
       // Parameter name definition
       #parameterDefinition.parameterNameString := 'VEL';
       #parameterDefinition.parameterNameNumber := -1;

       // Matching to PathData
       #parameterDefinition.followingValues[1].cmdParameters.pathDynamics.velocity := TRUE;

       // Priorities
       #parameterDefinition.priorities.cmdParameters.pathDynamics.velocity := "LKINLANG_PRIO_DEFINED";

       // Properties
       #parameterDefinition.properties := "LKINLANG_PRG_MODAL" + "LKINLANG_EQUATION";

       // Valid counts per line
       #parameterDefinition.validCountPerLine := 1;
       // ========================================================================================================
